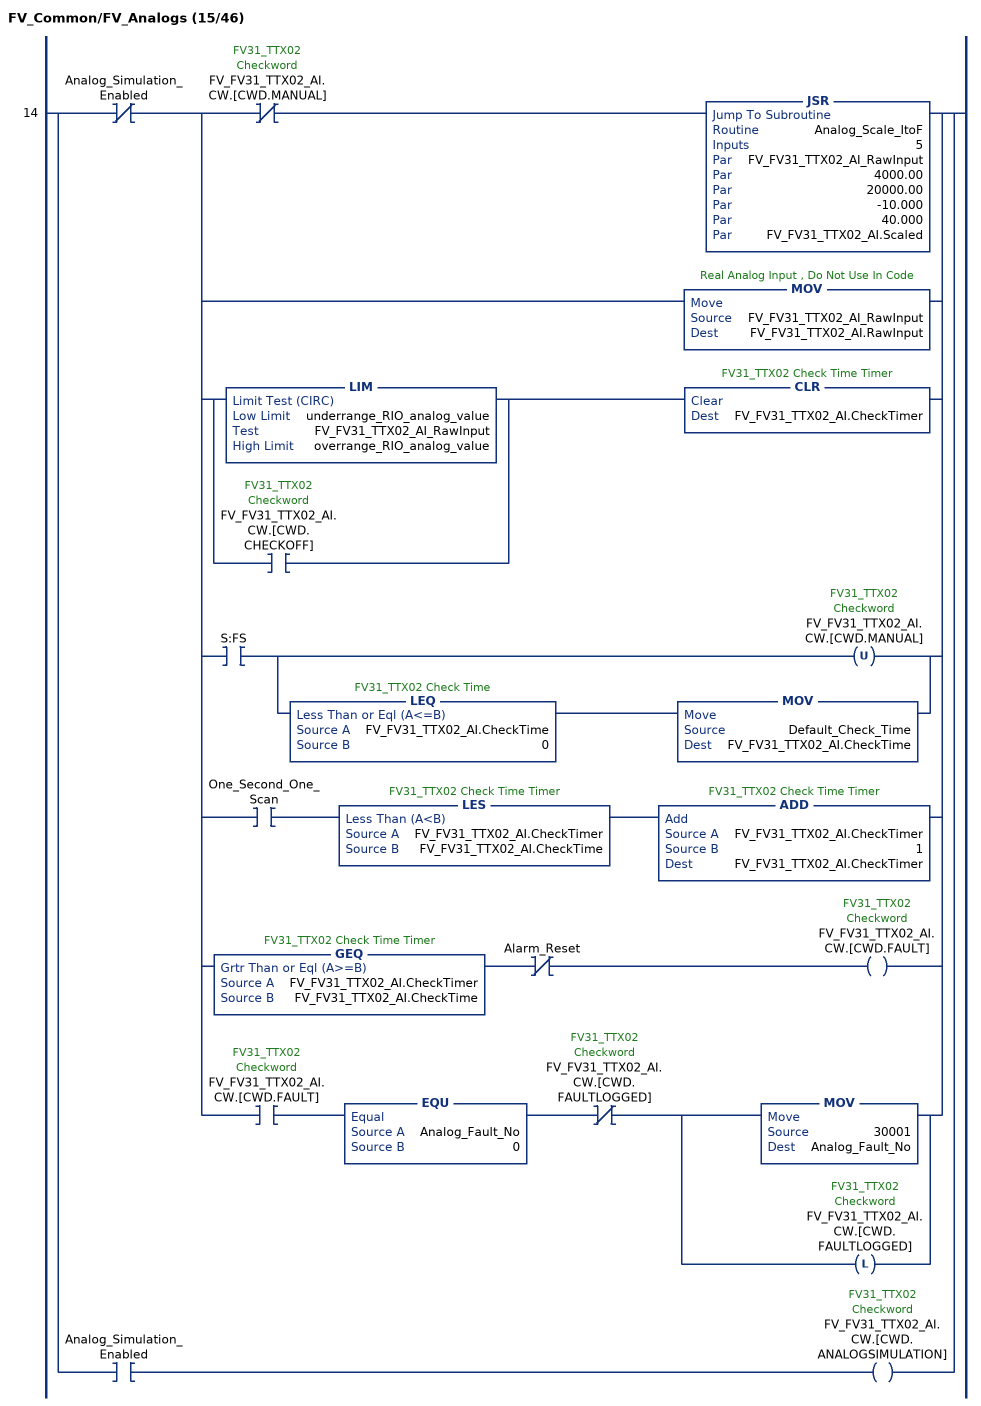
   14: [XIO(Analog_Simulation_Enabled) [XIO(FV_FV31_TTX02_AI.CW.[CWD.MANUAL]) JSR(Analog_Scale_ItoF,5,FV_FV31_TTX02_AI_RawInput,4000.00,20000.00,-10.000,40.000,FV_FV31_TTX02_AI.Scaled) ,MOV(FV_FV31_TTX02_AI_RawInput,FV_FV31_TTX02_AI.RawInput) ,[LIM(underrange_RIO_analog_value,FV_FV31_TTX02_AI_RawInput,overrange_RIO_analog_value) ,XIC(FV_FV31_TTX02_AI.CW.[CWD.CHECKOFF]) ] CLR(FV_FV31_TTX02_AI.CheckTimer) ,XIC(S:FS) [OTU(FV_FV31_TTX02_AI.CW.[CWD.MANUAL]) ,LEQ(FV_FV31_TTX02_AI.CheckTime,0) MOV(Default_Check_Time,FV_FV31_TTX02_AI.CheckTime) ] ,XIC(One_Second_One_Scan) LES(FV_FV31_TTX02_AI.CheckTimer,FV_FV31_TTX02_AI.CheckTime) ADD(FV_FV31_TTX02_AI.CheckTimer,1,FV_FV31_TTX02_AI.CheckTimer) ,GEQ(FV_FV31_TTX02_AI.CheckTimer,FV_FV31_TTX02_AI.CheckTime) XIO(Alarm_Reset) OTE(FV_FV31_TTX02_AI.CW.[CWD.FAULT]) ,XIC(FV_FV31_TTX02_AI.CW.[CWD.FAULT]) EQU(Analog_Fault_No,0) XIO(FV_FV31_TTX02_AI.CW.[CWD.FAULTLOGGED]) [MOV(30001,Analog_Fault_No) ,OTL(FV_FV31_TTX02_AI.CW.[CWD.FAULTLOGGED]) ] ] ,XIC(Analog_Simulation_Enabled) OTE(FV_FV31_TTX02_AI.CW.[CWD.ANALOGSIMULATION]) ];
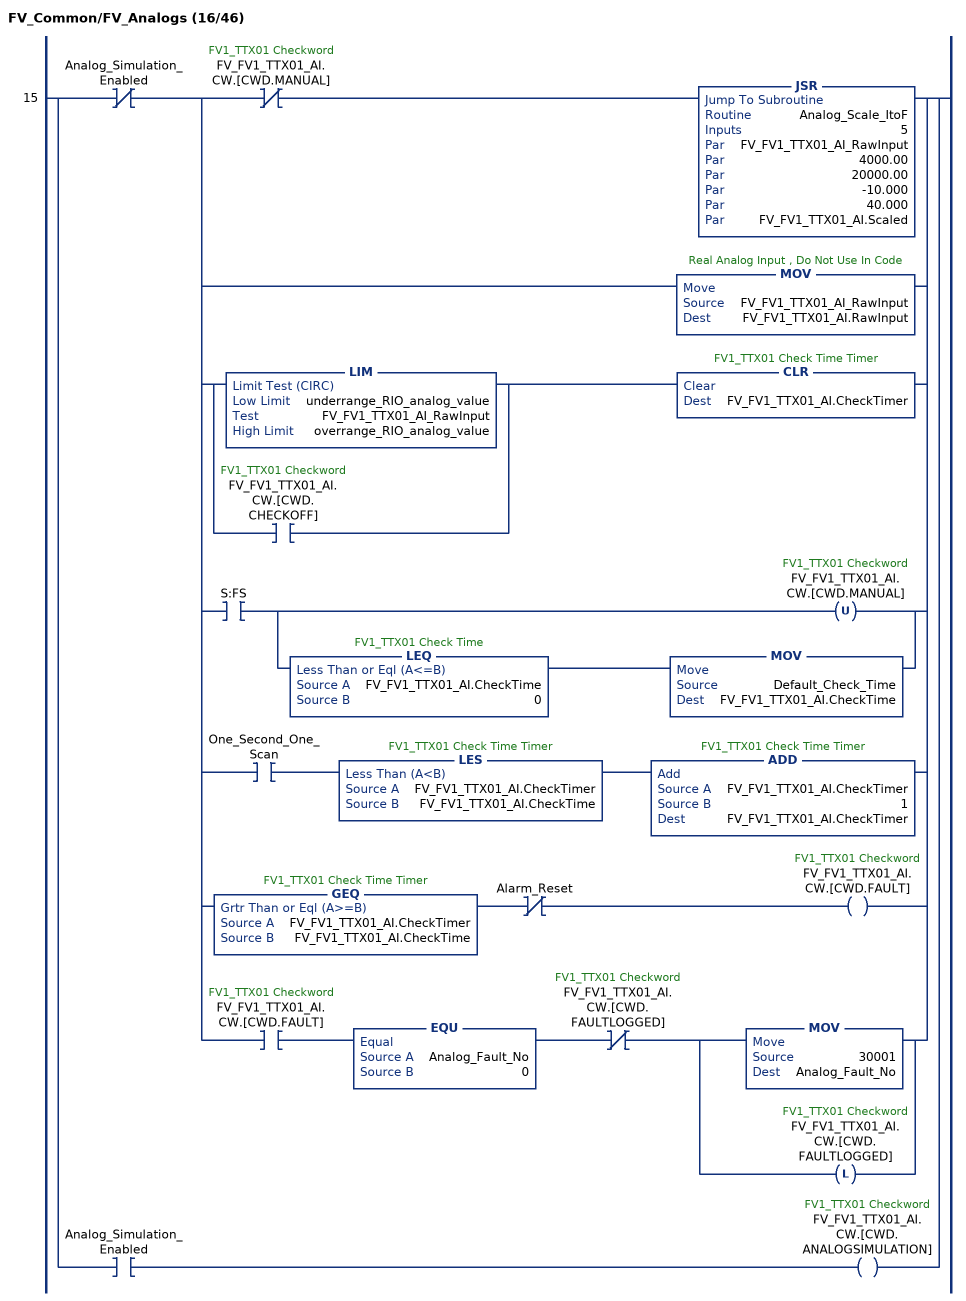
   15: [XIO(Analog_Simulation_Enabled) [XIO(FV_FV1_TTX01_AI.CW.[CWD.MANUAL]) JSR(Analog_Scale_ItoF,5,FV_FV1_TTX01_AI_RawInput,4000.00,20000.00,-10.000,40.000,FV_FV1_TTX01_AI.Scaled) ,MOV(FV_FV1_TTX01_AI_RawInput,FV_FV1_TTX01_AI.RawInput) ,[LIM(underrange_RIO_analog_value,FV_FV1_TTX01_AI_RawInput,overrange_RIO_analog_value) ,XIC(FV_FV1_TTX01_AI.CW.[CWD.CHECKOFF]) ] CLR(FV_FV1_TTX01_AI.CheckTimer) ,XIC(S:FS) [OTU(FV_FV1_TTX01_AI.CW.[CWD.MANUAL]) ,LEQ(FV_FV1_TTX01_AI.CheckTime,0) MOV(Default_Check_Time,FV_FV1_TTX01_AI.CheckTime) ] ,XIC(One_Second_One_Scan) LES(FV_FV1_TTX01_AI.CheckTimer,FV_FV1_TTX01_AI.CheckTime) ADD(FV_FV1_TTX01_AI.CheckTimer,1,FV_FV1_TTX01_AI.CheckTimer) ,GEQ(FV_FV1_TTX01_AI.CheckTimer,FV_FV1_TTX01_AI.CheckTime) XIO(Alarm_Reset) OTE(FV_FV1_TTX01_AI.CW.[CWD.FAULT]) ,XIC(FV_FV1_TTX01_AI.CW.[CWD.FAULT]) EQU(Analog_Fault_No,0) XIO(FV_FV1_TTX01_AI.CW.[CWD.FAULTLOGGED]) [MOV(30001,Analog_Fault_No) ,OTL(FV_FV1_TTX01_AI.CW.[CWD.FAULTLOGGED]) ] ] ,XIC(Analog_Simulation_Enabled) OTE(FV_FV1_TTX01_AI.CW.[CWD.ANALOGSIMULATION]) ];
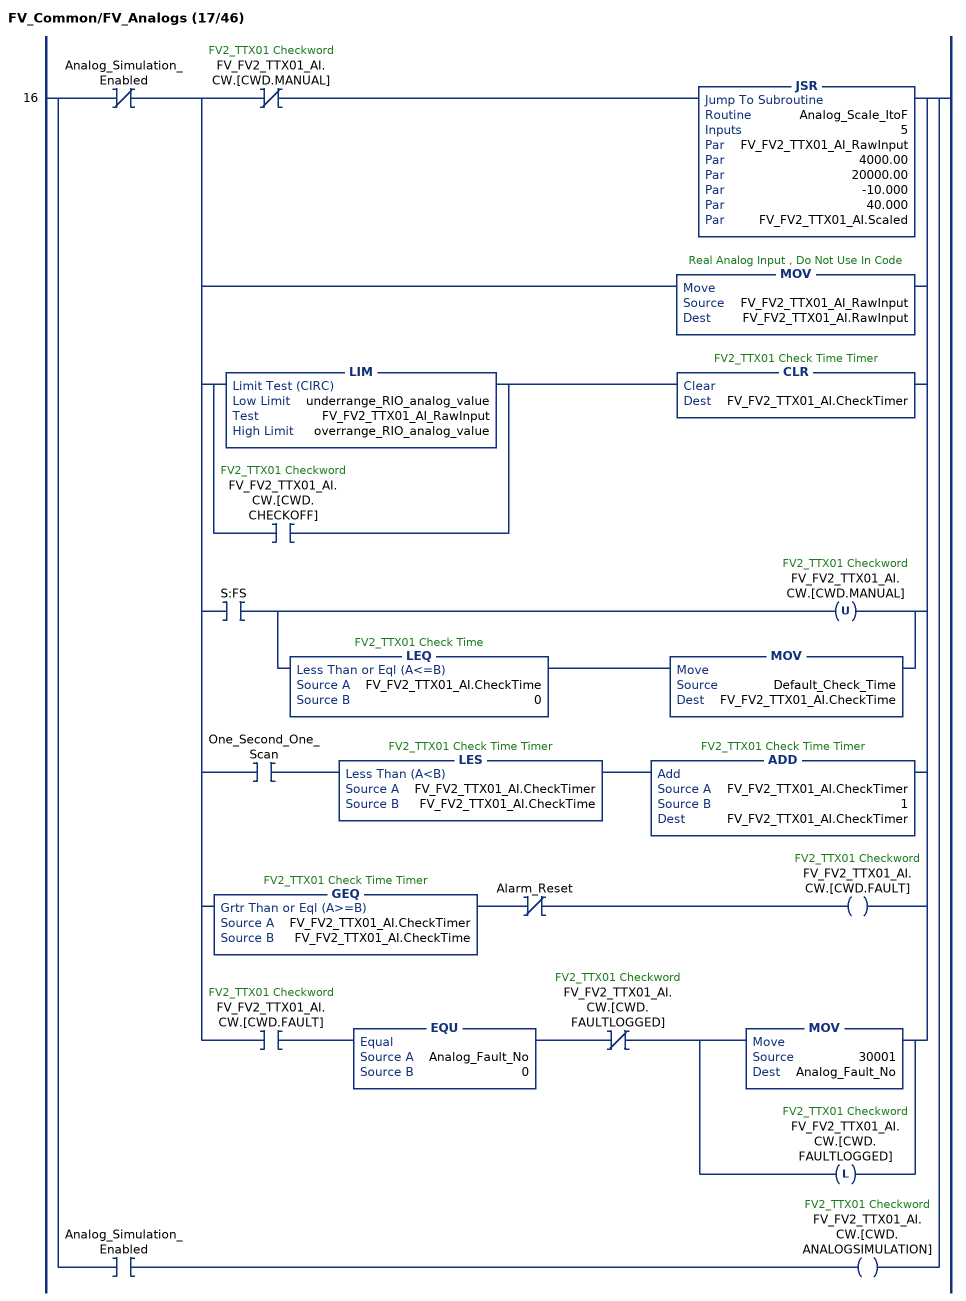
   16: [XIO(Analog_Simulation_Enabled) [XIO(FV_FV2_TTX01_AI.CW.[CWD.MANUAL]) JSR(Analog_Scale_ItoF,5,FV_FV2_TTX01_AI_RawInput,4000.00,20000.00,-10.000,40.000,FV_FV2_TTX01_AI.Scaled) ,MOV(FV_FV2_TTX01_AI_RawInput,FV_FV2_TTX01_AI.RawInput) ,[LIM(underrange_RIO_analog_value,FV_FV2_TTX01_AI_RawInput,overrange_RIO_analog_value) ,XIC(FV_FV2_TTX01_AI.CW.[CWD.CHECKOFF]) ] CLR(FV_FV2_TTX01_AI.CheckTimer) ,XIC(S:FS) [OTU(FV_FV2_TTX01_AI.CW.[CWD.MANUAL]) ,LEQ(FV_FV2_TTX01_AI.CheckTime,0) MOV(Default_Check_Time,FV_FV2_TTX01_AI.CheckTime) ] ,XIC(One_Second_One_Scan) LES(FV_FV2_TTX01_AI.CheckTimer,FV_FV2_TTX01_AI.CheckTime) ADD(FV_FV2_TTX01_AI.CheckTimer,1,FV_FV2_TTX01_AI.CheckTimer) ,GEQ(FV_FV2_TTX01_AI.CheckTimer,FV_FV2_TTX01_AI.CheckTime) XIO(Alarm_Reset) OTE(FV_FV2_TTX01_AI.CW.[CWD.FAULT]) ,XIC(FV_FV2_TTX01_AI.CW.[CWD.FAULT]) EQU(Analog_Fault_No,0) XIO(FV_FV2_TTX01_AI.CW.[CWD.FAULTLOGGED]) [MOV(30001,Analog_Fault_No) ,OTL(FV_FV2_TTX01_AI.CW.[CWD.FAULTLOGGED]) ] ] ,XIC(Analog_Simulation_Enabled) OTE(FV_FV2_TTX01_AI.CW.[CWD.ANALOGSIMULATION]) ];
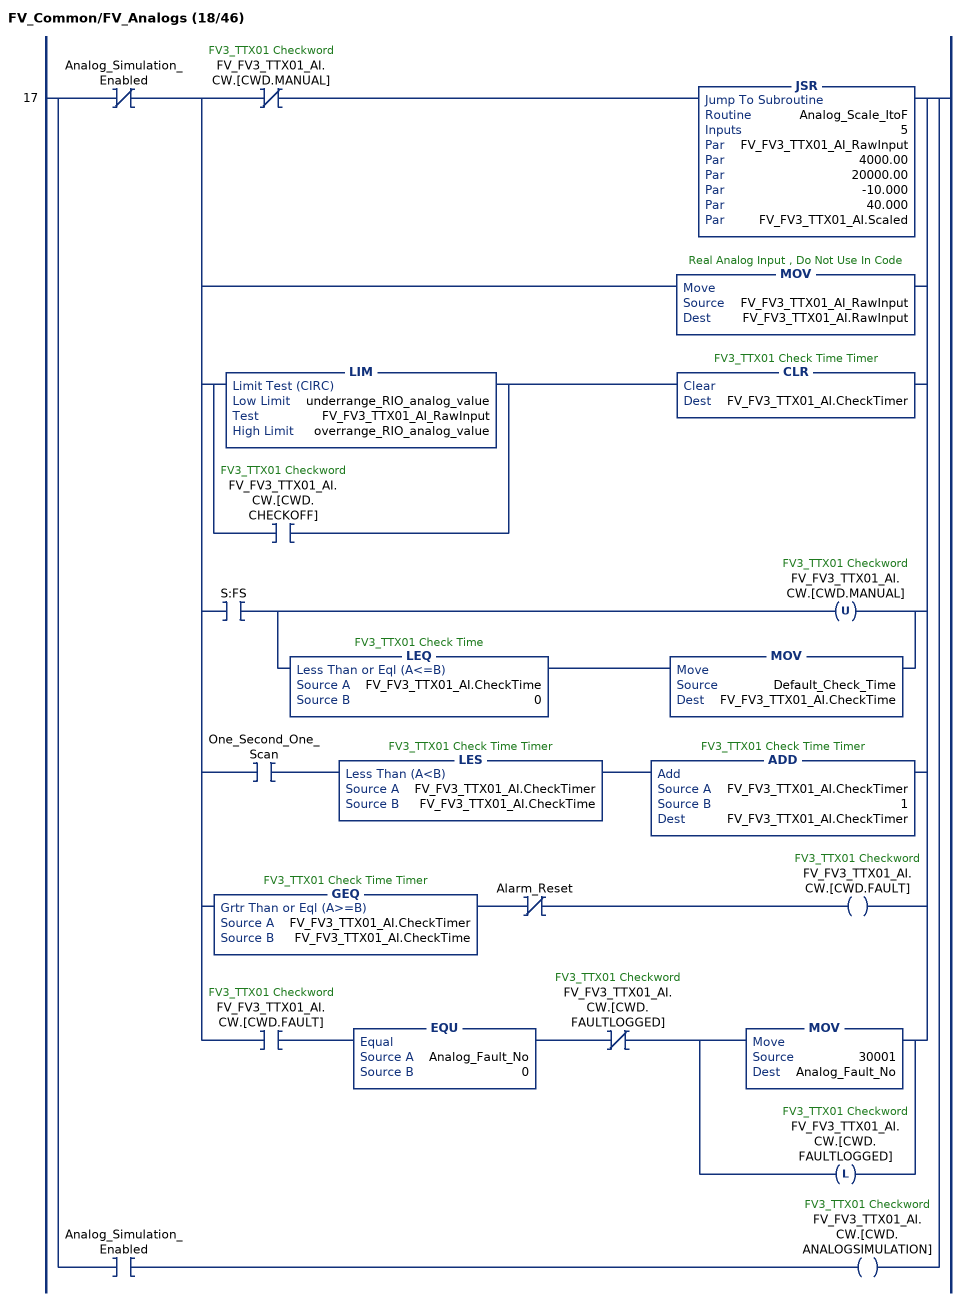
   17: [XIO(Analog_Simulation_Enabled) [XIO(FV_FV3_TTX01_AI.CW.[CWD.MANUAL]) JSR(Analog_Scale_ItoF,5,FV_FV3_TTX01_AI_RawInput,4000.00,20000.00,-10.000,40.000,FV_FV3_TTX01_AI.Scaled) ,MOV(FV_FV3_TTX01_AI_RawInput,FV_FV3_TTX01_AI.RawInput) ,[LIM(underrange_RIO_analog_value,FV_FV3_TTX01_AI_RawInput,overrange_RIO_analog_value) ,XIC(FV_FV3_TTX01_AI.CW.[CWD.CHECKOFF]) ] CLR(FV_FV3_TTX01_AI.CheckTimer) ,XIC(S:FS) [OTU(FV_FV3_TTX01_AI.CW.[CWD.MANUAL]) ,LEQ(FV_FV3_TTX01_AI.CheckTime,0) MOV(Default_Check_Time,FV_FV3_TTX01_AI.CheckTime) ] ,XIC(One_Second_One_Scan) LES(FV_FV3_TTX01_AI.CheckTimer,FV_FV3_TTX01_AI.CheckTime) ADD(FV_FV3_TTX01_AI.CheckTimer,1,FV_FV3_TTX01_AI.CheckTimer) ,GEQ(FV_FV3_TTX01_AI.CheckTimer,FV_FV3_TTX01_AI.CheckTime) XIO(Alarm_Reset) OTE(FV_FV3_TTX01_AI.CW.[CWD.FAULT]) ,XIC(FV_FV3_TTX01_AI.CW.[CWD.FAULT]) EQU(Analog_Fault_No,0) XIO(FV_FV3_TTX01_AI.CW.[CWD.FAULTLOGGED]) [MOV(30001,Analog_Fault_No) ,OTL(FV_FV3_TTX01_AI.CW.[CWD.FAULTLOGGED]) ] ] ,XIC(Analog_Simulation_Enabled) OTE(FV_FV3_TTX01_AI.CW.[CWD.ANALOGSIMULATION]) ];
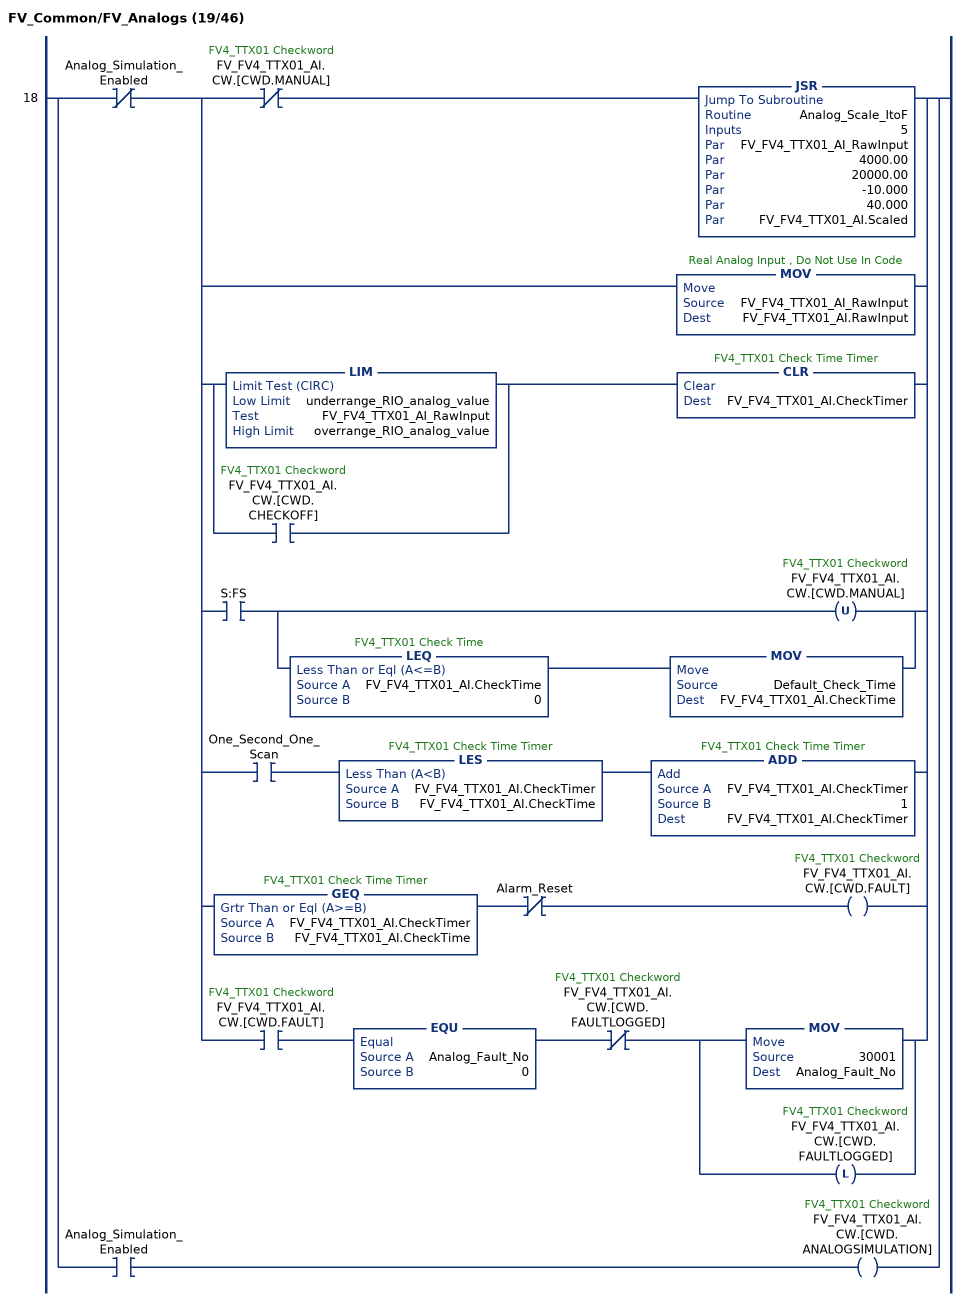
   18: [XIO(Analog_Simulation_Enabled) [XIO(FV_FV4_TTX01_AI.CW.[CWD.MANUAL]) JSR(Analog_Scale_ItoF,5,FV_FV4_TTX01_AI_RawInput,4000.00,20000.00,-10.000,40.000,FV_FV4_TTX01_AI.Scaled) ,MOV(FV_FV4_TTX01_AI_RawInput,FV_FV4_TTX01_AI.RawInput) ,[LIM(underrange_RIO_analog_value,FV_FV4_TTX01_AI_RawInput,overrange_RIO_analog_value) ,XIC(FV_FV4_TTX01_AI.CW.[CWD.CHECKOFF]) ] CLR(FV_FV4_TTX01_AI.CheckTimer) ,XIC(S:FS) [OTU(FV_FV4_TTX01_AI.CW.[CWD.MANUAL]) ,LEQ(FV_FV4_TTX01_AI.CheckTime,0) MOV(Default_Check_Time,FV_FV4_TTX01_AI.CheckTime) ] ,XIC(One_Second_One_Scan) LES(FV_FV4_TTX01_AI.CheckTimer,FV_FV4_TTX01_AI.CheckTime) ADD(FV_FV4_TTX01_AI.CheckTimer,1,FV_FV4_TTX01_AI.CheckTimer) ,GEQ(FV_FV4_TTX01_AI.CheckTimer,FV_FV4_TTX01_AI.CheckTime) XIO(Alarm_Reset) OTE(FV_FV4_TTX01_AI.CW.[CWD.FAULT]) ,XIC(FV_FV4_TTX01_AI.CW.[CWD.FAULT]) EQU(Analog_Fault_No,0) XIO(FV_FV4_TTX01_AI.CW.[CWD.FAULTLOGGED]) [MOV(30001,Analog_Fault_No) ,OTL(FV_FV4_TTX01_AI.CW.[CWD.FAULTLOGGED]) ] ] ,XIC(Analog_Simulation_Enabled) OTE(FV_FV4_TTX01_AI.CW.[CWD.ANALOGSIMULATION]) ];
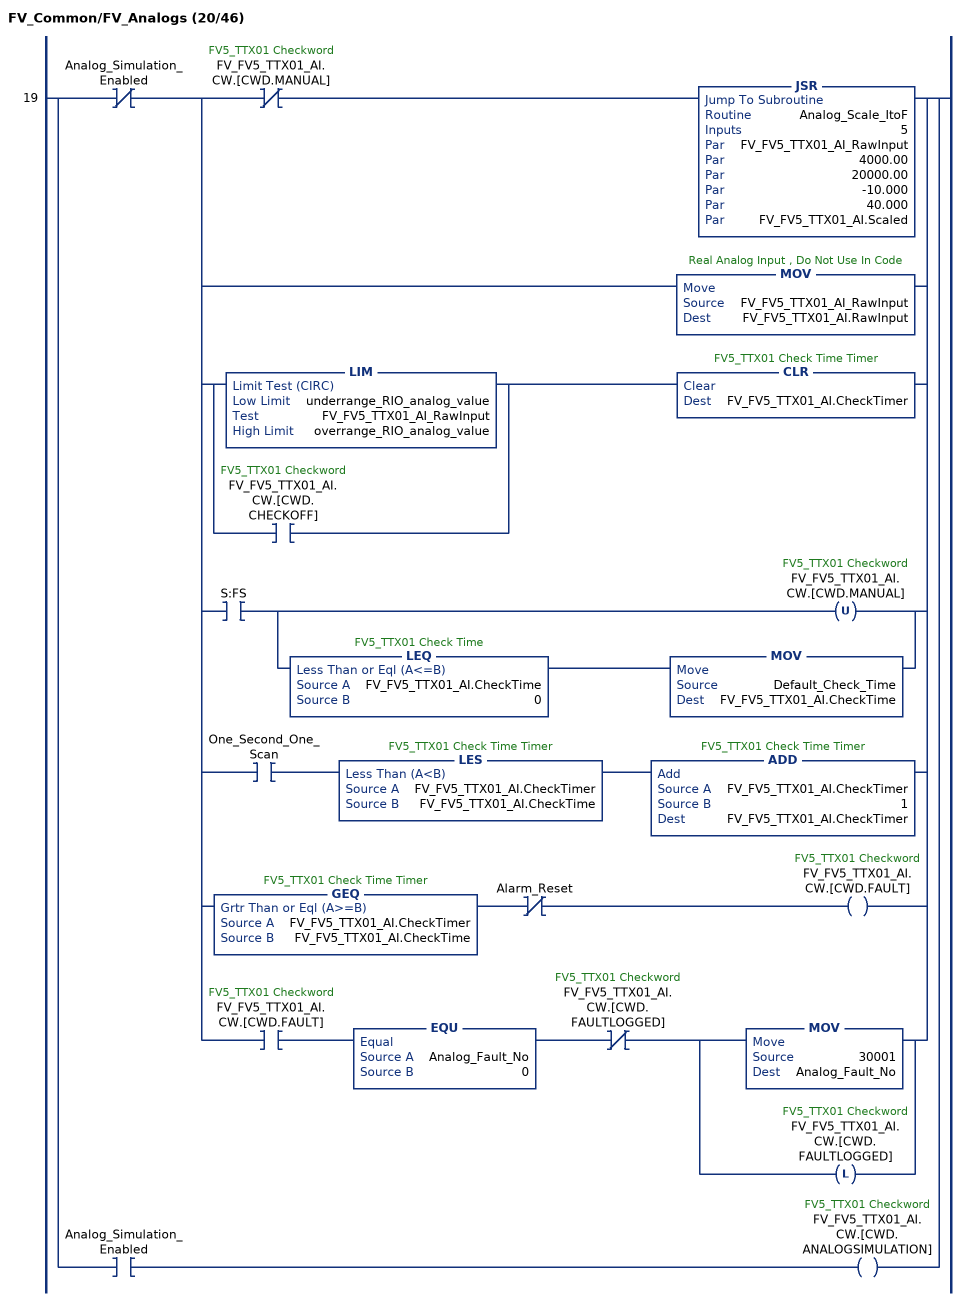
   19: [XIO(Analog_Simulation_Enabled) [XIO(FV_FV5_TTX01_AI.CW.[CWD.MANUAL]) JSR(Analog_Scale_ItoF,5,FV_FV5_TTX01_AI_RawInput,4000.00,20000.00,-10.000,40.000,FV_FV5_TTX01_AI.Scaled) ,MOV(FV_FV5_TTX01_AI_RawInput,FV_FV5_TTX01_AI.RawInput) ,[LIM(underrange_RIO_analog_value,FV_FV5_TTX01_AI_RawInput,overrange_RIO_analog_value) ,XIC(FV_FV5_TTX01_AI.CW.[CWD.CHECKOFF]) ] CLR(FV_FV5_TTX01_AI.CheckTimer) ,XIC(S:FS) [OTU(FV_FV5_TTX01_AI.CW.[CWD.MANUAL]) ,LEQ(FV_FV5_TTX01_AI.CheckTime,0) MOV(Default_Check_Time,FV_FV5_TTX01_AI.CheckTime) ] ,XIC(One_Second_One_Scan) LES(FV_FV5_TTX01_AI.CheckTimer,FV_FV5_TTX01_AI.CheckTime) ADD(FV_FV5_TTX01_AI.CheckTimer,1,FV_FV5_TTX01_AI.CheckTimer) ,GEQ(FV_FV5_TTX01_AI.CheckTimer,FV_FV5_TTX01_AI.CheckTime) XIO(Alarm_Reset) OTE(FV_FV5_TTX01_AI.CW.[CWD.FAULT]) ,XIC(FV_FV5_TTX01_AI.CW.[CWD.FAULT]) EQU(Analog_Fault_No,0) XIO(FV_FV5_TTX01_AI.CW.[CWD.FAULTLOGGED]) [MOV(30001,Analog_Fault_No) ,OTL(FV_FV5_TTX01_AI.CW.[CWD.FAULTLOGGED]) ] ] ,XIC(Analog_Simulation_Enabled) OTE(FV_FV5_TTX01_AI.CW.[CWD.ANALOGSIMULATION]) ];
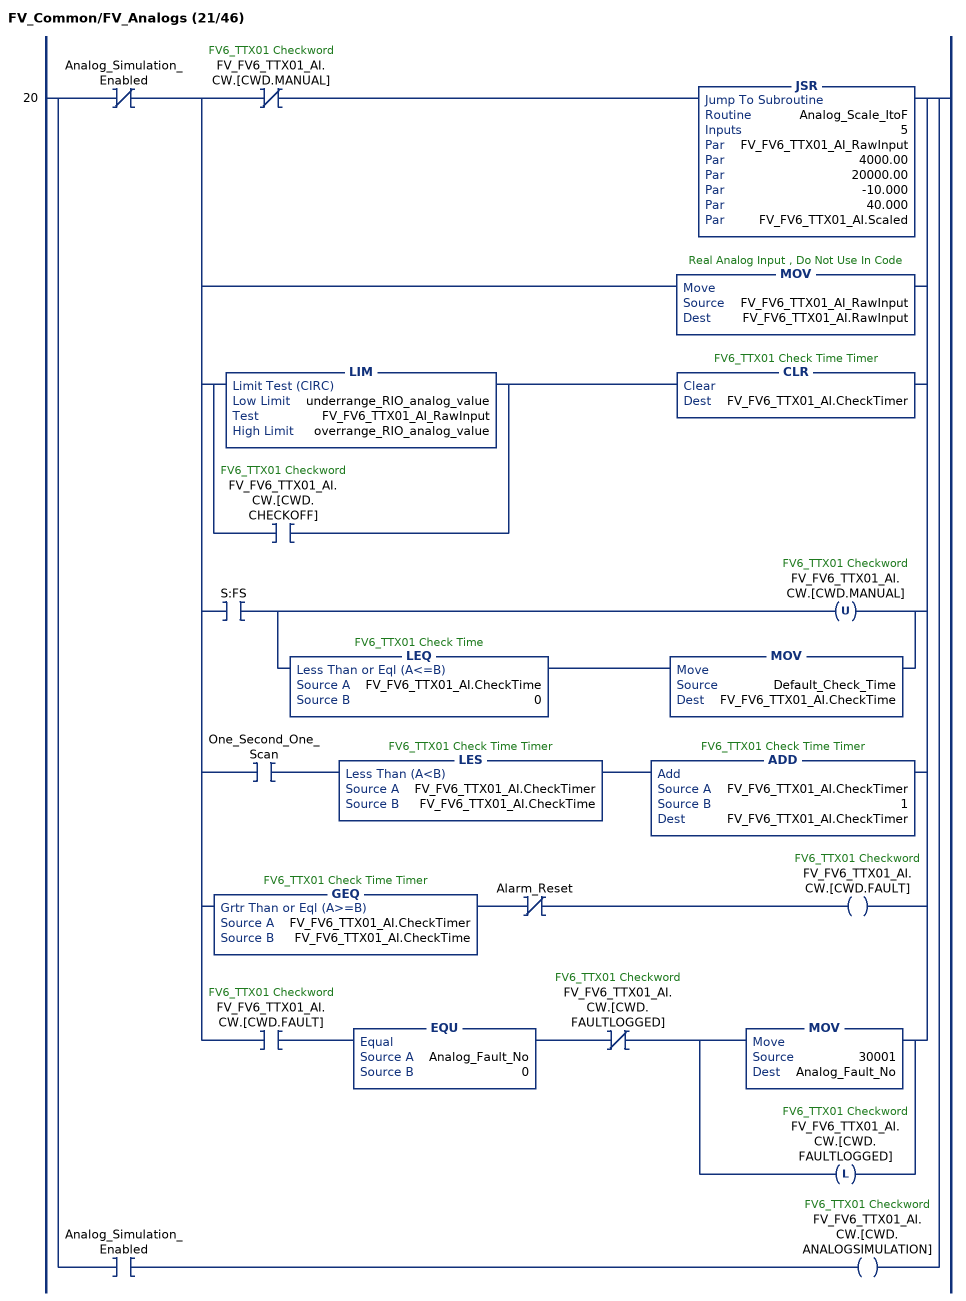
   20: [XIO(Analog_Simulation_Enabled) [XIO(FV_FV6_TTX01_AI.CW.[CWD.MANUAL]) JSR(Analog_Scale_ItoF,5,FV_FV6_TTX01_AI_RawInput,4000.00,20000.00,-10.000,40.000,FV_FV6_TTX01_AI.Scaled) ,MOV(FV_FV6_TTX01_AI_RawInput,FV_FV6_TTX01_AI.RawInput) ,[LIM(underrange_RIO_analog_value,FV_FV6_TTX01_AI_RawInput,overrange_RIO_analog_value) ,XIC(FV_FV6_TTX01_AI.CW.[CWD.CHECKOFF]) ] CLR(FV_FV6_TTX01_AI.CheckTimer) ,XIC(S:FS) [OTU(FV_FV6_TTX01_AI.CW.[CWD.MANUAL]) ,LEQ(FV_FV6_TTX01_AI.CheckTime,0) MOV(Default_Check_Time,FV_FV6_TTX01_AI.CheckTime) ] ,XIC(One_Second_One_Scan) LES(FV_FV6_TTX01_AI.CheckTimer,FV_FV6_TTX01_AI.CheckTime) ADD(FV_FV6_TTX01_AI.CheckTimer,1,FV_FV6_TTX01_AI.CheckTimer) ,GEQ(FV_FV6_TTX01_AI.CheckTimer,FV_FV6_TTX01_AI.CheckTime) XIO(Alarm_Reset) OTE(FV_FV6_TTX01_AI.CW.[CWD.FAULT]) ,XIC(FV_FV6_TTX01_AI.CW.[CWD.FAULT]) EQU(Analog_Fault_No,0) XIO(FV_FV6_TTX01_AI.CW.[CWD.FAULTLOGGED]) [MOV(30001,Analog_Fault_No) ,OTL(FV_FV6_TTX01_AI.CW.[CWD.FAULTLOGGED]) ] ] ,XIC(Analog_Simulation_Enabled) OTE(FV_FV6_TTX01_AI.CW.[CWD.ANALOGSIMULATION]) ];
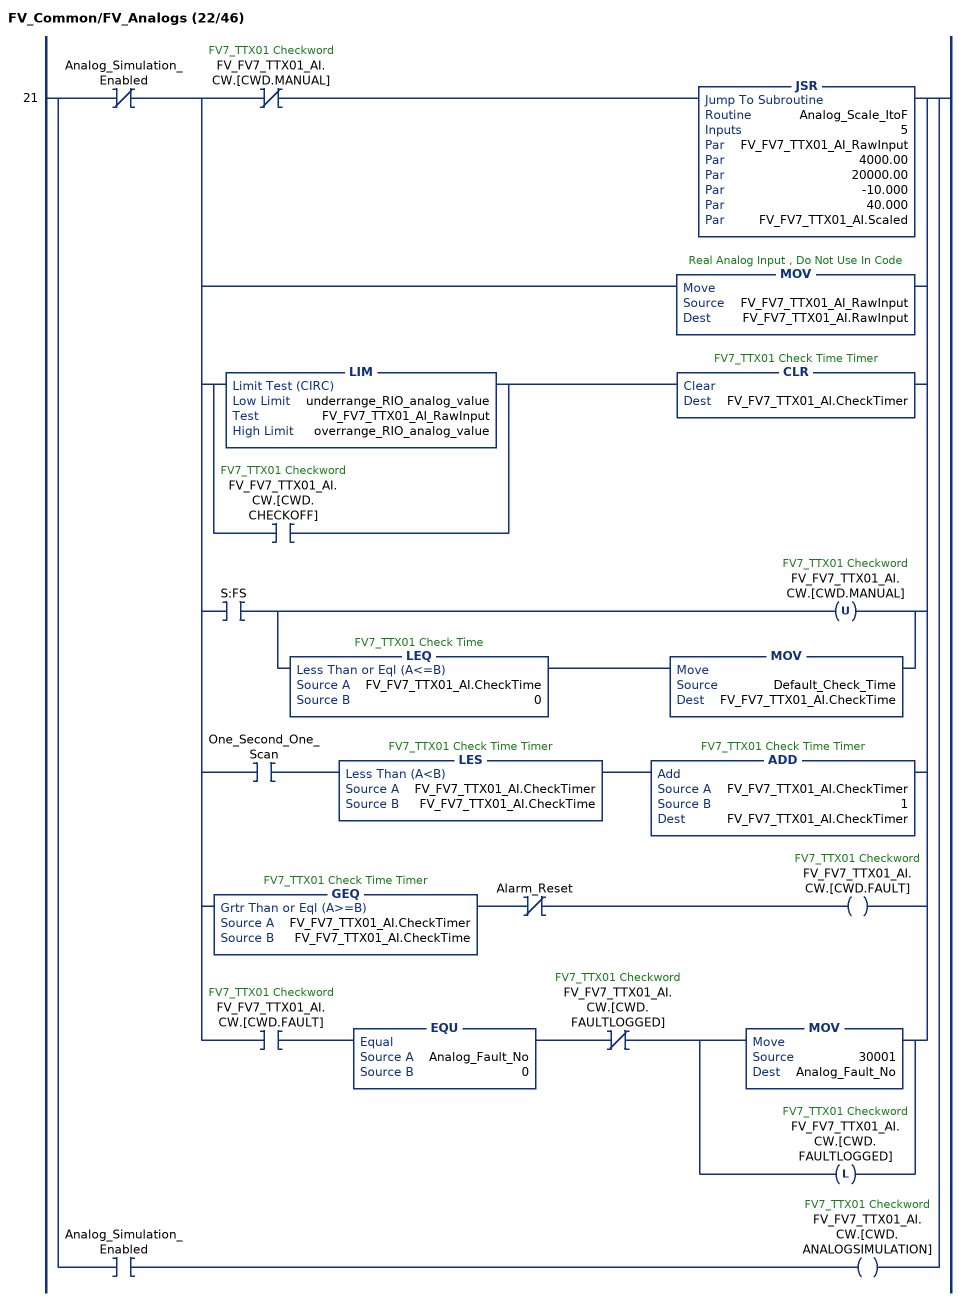
   21: [XIO(Analog_Simulation_Enabled) [XIO(FV_FV7_TTX01_AI.CW.[CWD.MANUAL]) JSR(Analog_Scale_ItoF,5,FV_FV7_TTX01_AI_RawInput,4000.00,20000.00,-10.000,40.000,FV_FV7_TTX01_AI.Scaled) ,MOV(FV_FV7_TTX01_AI_RawInput,FV_FV7_TTX01_AI.RawInput) ,[LIM(underrange_RIO_analog_value,FV_FV7_TTX01_AI_RawInput,overrange_RIO_analog_value) ,XIC(FV_FV7_TTX01_AI.CW.[CWD.CHECKOFF]) ] CLR(FV_FV7_TTX01_AI.CheckTimer) ,XIC(S:FS) [OTU(FV_FV7_TTX01_AI.CW.[CWD.MANUAL]) ,LEQ(FV_FV7_TTX01_AI.CheckTime,0) MOV(Default_Check_Time,FV_FV7_TTX01_AI.CheckTime) ] ,XIC(One_Second_One_Scan) LES(FV_FV7_TTX01_AI.CheckTimer,FV_FV7_TTX01_AI.CheckTime) ADD(FV_FV7_TTX01_AI.CheckTimer,1,FV_FV7_TTX01_AI.CheckTimer) ,GEQ(FV_FV7_TTX01_AI.CheckTimer,FV_FV7_TTX01_AI.CheckTime) XIO(Alarm_Reset) OTE(FV_FV7_TTX01_AI.CW.[CWD.FAULT]) ,XIC(FV_FV7_TTX01_AI.CW.[CWD.FAULT]) EQU(Analog_Fault_No,0) XIO(FV_FV7_TTX01_AI.CW.[CWD.FAULTLOGGED]) [MOV(30001,Analog_Fault_No) ,OTL(FV_FV7_TTX01_AI.CW.[CWD.FAULTLOGGED]) ] ] ,XIC(Analog_Simulation_Enabled) OTE(FV_FV7_TTX01_AI.CW.[CWD.ANALOGSIMULATION]) ];
